   "Carrier_78_SpareSafetyInput(2_3)" AT %I4264.3 : Bool;   // SPARE SAFETY INPUT
   "Carrier_78_SpareSafetyInput(2_4)" AT %I4264.4 : Bool;   // SPARE SAFETY INPUT
   "Carrier_78_SpareSafetyInput(2_5)" AT %I4264.5 : Bool;   // SPARE SAFETY INPUT
   "Carrier_78_SpareSafetyInput(2_6)" AT %I4264.6 : Bool;   // SPARE SAFETY INPUT
   "Carrier_78_SpareSafetyInput(2_7)" AT %I4264.7 : Bool;   // SPARE SAFETY INPUT
   "Carrier_78_Slot3_SafetyOutput" AT %IW4265 : Word;   // SLOT 3 SAFETY OUTPUT WORD
   "Carrier_78_Crash_Detect_OK" AT %I4265.0 : Bool;   // CARRIER CRASH DETECT
   "Carrier_78_SpareSafetyOutput(3_1)" AT %I4265.1 : Bool;   // SPARE SAFETY OUTPUT
   "Carrier_78_SpareSafetyOutput(3_2)" AT %I4265.2 : Bool;   // SPARE SAFETY OUTPUT
   "Carrier_78_SpareSafetyOutput(3_3)" AT %I4265.3 : Bool;   // SPARE SAFETY OUTPUT
   "Carrier_78_SpareSafetyOutput(3_4)" AT %I4265.4 : Bool;   // SPARE SAFETY OUTPUT
   "Carrier_78_SpareSafetyOutput(3_5)" AT %I4265.5 : Bool;   // SPARE SAFETY OUTPUT
   "Carrier_78_SpareSafetyOutput(3_6)" AT %I4265.6 : Bool;   // SPARE SAFETY OUTPUT
   "Carrier_78_SpareSafetyOutput(3_7)" AT %I4265.7 : Bool;   // SPARE SAFETY OUTPUT
   "Carrier_78_Slot4_Input" AT %IW4266 : Word;   // SLOT 4 INPUT WORD
   "Carrier_78_480VPowerOn_MDCB1" AT %I4266.0 : Bool;   // 480 VAC POWER ON MDCB 1
   "Carrier_78_SpareInput(4_1)" AT %I4266.1 : Bool;   // SPARE INPUT
   "Carrier_78_SpareInput(4_2)" AT %I4266.2 : Bool;   // SPARE INPUT
   "Carrier_78_SitopSelectStatus" AT %I4266.3 : Bool;   // SITOP SELECT STATUS
   "Carrier_78_DCsupplyOnPSCB2" AT %I4266.4 : Bool;   // DC SUPPLY ON PSCB 2
   "Carrier_78_SpareInput(4_5)" AT %I4266.5 : Bool;   // SPARE INPUT
   "Carrier_78_SpareInput(4_6)" AT %I4266.6 : Bool;   // SPARE INPUT
   "Carrier_78_SpareInput(4_7)" AT %I4266.7 : Bool;   // SPARE INPUT
   "Carrier_78_PB1_ProdHoldLH" AT %I4267.0 : Bool;   // PB 1 PRODUCTION HOLD LH
   "Carrier_78_PB2_ResetLH" AT %I4267.1 : Bool;   // PB 2 RESET LH
   "Carrier_78_PB3_ProdHoldRH" AT %I4267.2 : Bool;   // PB 3 PRODUCTION HOLD RH
   "Carrier_78_PB4_ResetRH" AT %I4267.3 : Bool;   // PB 4 RESET RH
   "Carrier_78_SpareInput(4_14)" AT %I4267.4 : Bool;   // SPARE INPUT
   "Carrier_78_SpareInput(4_15)" AT %I4267.5 : Bool;   // SPARE INPUT
   "Carrier_78_SpareInput(4_16)" AT %I4267.6 : Bool;   // SPARE INPUT
   "Carrier_78_SpareInput(4_17)" AT %I4267.7 : Bool;   // SPARE INPUT
   "Carrier_78_Slot5_Output" AT %IW4268 : Word;   // SLOT 5 OUTPUT WORD
   "Carrier_78_IRD400_HMI_24VDC_ENABLE" AT %I4268.0 : Bool;   // IRD 400 PANEL HMI 24V DC POWER
   "Carrier_78_FaultLight_LH" AT %I4268.1 : Bool;   // FAULT LIGHT LH
   "Carrier_78_RunLight_LH" AT %I4268.2 : Bool;   // RUN LIGHT LH
   "Carrier_78_FaultLight_RH" AT %I4268.3 : Bool;   // FAULT LIGHT RH
   "Carrier_78_RunLight_RH" AT %I4268.4 : Bool;   // RUN LIGHT RH
   "Carrier_78_SpareOutput(5_5)" AT %I4268.5 : Bool;   // SPARE OUTPUT
   "Carrier_78_SpareOutput(5_6)" AT %I4268.6 : Bool;   // SPARE OUTPUT
   "Carrier_78_SpareOutput(5_7)" AT %I4268.7 : Bool;   // SPARE OUTPUT
   "Carrier_78_ActualSpeed" AT %IW4270 : Word;   // ACTUAL SPEED
   "Carrier_78_CarrierDriveAlarm" AT %IW4272 : Word;   // CARRIER DRIVE ALARM
   "Carrier_78_CarrierDriveWarning" AT %IW4274 : Word;   // CARRIER DRIVE WARNING
   "Carrier_79_Status" AT %IW4300 : Word;   // CARRIER STATUS WORD
   "Carrier_79_Status.0" AT %I4300.0 : Bool;   // HEARTBEAT
   "Carrier_79_Status.1" AT %I4300.1 : Bool;   // MANUAL
   "Carrier_79_Status.2" AT %I4300.2 : Bool;   // IN_AUTO
   "Carrier_79_Status.3" AT %I4300.3 : Bool;   // POSITIONING_COMPLETE
   "Carrier_79_Status.4" AT %I4300.4 : Bool;   // PRODUCTION HOLD
   "Carrier_79_Status.5" AT %I4300.5 : Bool;   // CARRIER MOVING FORWARD
   "Carrier_79_Status.6" AT %I4300.6 : Bool;   // CARRIER MOVING REVERSE
   "Carrier_79_Status.7" AT %I4300.7 : Bool;   // CARRIER FAULT
   "Carrier_79_Status.8" AT %I4301.0 : Bool;   // CRASH DETECT TRIPPED
   "Carrier_79_Status.9" AT %I4301.1 : Bool;
   "Carrier_79_Status.10" AT %I4301.2 : Bool;
   "Carrier_79_Status.11" AT %I4301.3 : Bool;
   "Carrier_79_Status.12" AT %I4301.4 : Bool;
   "Carrier_79_Status.13" AT %I4301.5 : Bool;
   "Carrier_79_Status.14" AT %I4301.6 : Bool;
   "Carrier_79_Status.15" AT %I4301.7 : Bool;
   "Carrier_79_SDCFaultCode" AT %IW4302 : Word;   // SDC FAULT CODE
   "Carrier_79_CarrierPosition" AT %ID4304 : DWord;   // CARRIER POSITION
   "Carrier_79_CarrierNumber" AT %IW4308 : Word;   // CARRIER NUMBER
   "Carrier_79_G120DControlWord" AT %IW4310 : Word;   // G120D_STW1_CONTROL
   "Carrier_79_G120DControlWord.0" AT %I4310.0 : Bool;   // Bit_00_ON
   "Carrier_79_G120DControlWord.1" AT %I4310.1 : Bool;   // Bit_01_AUS2_INH
   "Carrier_79_G120DControlWord.2" AT %I4310.2 : Bool;   // Bit_02_AUS3_STOP
   "Carrier_79_G120DControlWord.3" AT %I4310.3 : Bool;   // Bit_03_EN
   "Carrier_79_G120DControlWord.4" AT %I4310.4 : Bool;   // Bit_04_EN_RAMP
   "Carrier_79_G120DControlWord.5" AT %I4310.5 : Bool;   // Bit_05_START_RAMP
   "Carrier_79_G120DControlWord.6" AT %I4310.6 : Bool;   // Bit_06_SETPOINT
   "Carrier_79_G120DControlWord.7" AT %I4310.7 : Bool;   // Bit_07_RESET
   "Carrier_79_G120DControlWord.8" AT %I4311.0 : Bool;   // Bit_08_JOG_R
   "Carrier_79_G120DControlWord.9" AT %I4311.1 : Bool;   // Bit_09_JOG_L
   "Carrier_79_G120DControlWord.10" AT %I4311.2 : Bool;   // Bit_10_CONTR_PLC
   "Carrier_79_G120DControlWord.11" AT %I4311.3 : Bool;   // Bit_11_REVERSE
   "Carrier_79_G120DControlWord.12" AT %I4311.4 : Bool;   // Bit_12_BRAKE_RELEASE
   "Carrier_79_G120DControlWord.13" AT %I4311.5 : Bool;   // Bit_13_DDS
   "Carrier_79_G120DControlWord.14" AT %I4311.6 : Bool;   // Bit_14_DO0
   "Carrier_79_G120DControlWord.15" AT %I4311.7 : Bool;   // Bit_15_DO1
   "Carrier_79_G120DStatusWord" AT %IW4312 : Word;   // G120D_ZSW1_STATUS
   "Carrier_79_G120DStatusWord.0" AT %I4312.0 : Bool;   // Bit_00_READY_RUN
   "Carrier_79_G120DStatusWord.1" AT %I4312.1 : Bool;   // Bit_01_READY_ON
   "Carrier_79_G120DStatusWord.2" AT %I4312.2 : Bool;   // Bit_02_ENABLE
   "Carrier_79_G120DStatusWord.3" AT %I4312.3 : Bool;   // Bit_03_FAULT
   "Carrier_79_G120DStatusWord.4" AT %I4312.4 : Bool;   // Bit_04_OFF2
   "Carrier_79_G120DStatusWord.5" AT %I4312.5 : Bool;   // Bit_05_OFF3
   "Carrier_79_G120DStatusWord.6" AT %I4312.6 : Bool;   // Bit_06_LOCK_OUT
   "Carrier_79_G120DStatusWord.7" AT %I4312.7 : Bool;   // Bit_07_WARN
   "Carrier_79_G120DStatusWord.8" AT %I4313.0 : Bool;   // Bit_08_NO_DEVIATION
   "Carrier_79_G120DStatusWord.9" AT %I4313.1 : Bool;   // Bit_09_CONTR_PLC
   "Carrier_79_G120DStatusWord.10" AT %I4313.2 : Bool;   // Bit_10_F_MAX
   "Carrier_79_G120DStatusWord.11" AT %I4313.3 : Bool;   // Bit_11_LIMIT_REACHED
   "Carrier_79_G120DStatusWord.12" AT %I4313.4 : Bool;   // Bit_12_BRAKE_OPEN
   "Carrier_79_G120DStatusWord.13" AT %I4313.5 : Bool;   // Bit_13_NO_OVERTEMP
   "Carrier_79_G120DStatusWord.14" AT %I4313.6 : Bool;   // Bit_14_CW_CCW
   "Carrier_79_G120DStatusWord.15" AT %I4313.7 : Bool;   // Bit_15_OVERL
   "Carrier_79_Slot2_Input" AT %IW4314 : Word;   // SLOT 2 INPUT WORD
   "Carrier_79_CrashDetectSW" AT %I4314.0 : Bool;   // CRASH DETECT SW
   "Carrier_79_SpareSafetyInput(2_1)" AT %I4314.1 : Bool;   // SPARE SAFETY INPUT
   "Carrier_79_SpareSafetyInput(2_2)" AT %I4314.2 : Bool;   // SPARE SAFETY INPUT
   "Carrier_79_SpareSafetyInput(2_3)" AT %I4314.3 : Bool;   // SPARE SAFETY INPUT
   "Carrier_79_SpareSafetyInput(2_4)" AT %I4314.4 : Bool;   // SPARE SAFETY INPUT
   "Carrier_79_SpareSafetyInput(2_5)" AT %I4314.5 : Bool;   // SPARE SAFETY INPUT
   "Carrier_79_SpareSafetyInput(2_6)" AT %I4314.6 : Bool;   // SPARE SAFETY INPUT
   "Carrier_79_SpareSafetyInput(2_7)" AT %I4314.7 : Bool;   // SPARE SAFETY INPUT
   "Carrier_79_Slot3_SafetyOutput" AT %IW4315 : Word;   // SLOT 3 SAFETY OUTPUT WORD
   "Carrier_79_Crash_Detect_OK" AT %I4315.0 : Bool;   // CARRIER CRASH DETECT
   "Carrier_79_SpareSafetyOutput(3_1)" AT %I4315.1 : Bool;   // SPARE SAFETY OUTPUT
   "Carrier_79_SpareSafetyOutput(3_2)" AT %I4315.2 : Bool;   // SPARE SAFETY OUTPUT
   "Carrier_79_SpareSafetyOutput(3_3)" AT %I4315.3 : Bool;   // SPARE SAFETY OUTPUT
   "Carrier_79_SpareSafetyOutput(3_4)" AT %I4315.4 : Bool;   // SPARE SAFETY OUTPUT
   "Carrier_79_SpareSafetyOutput(3_5)" AT %I4315.5 : Bool;   // SPARE SAFETY OUTPUT
   "Carrier_79_SpareSafetyOutput(3_6)" AT %I4315.6 : Bool;   // SPARE SAFETY OUTPUT
   "Carrier_79_SpareSafetyOutput(3_7)" AT %I4315.7 : Bool;   // SPARE SAFETY OUTPUT
   "Carrier_79_Slot4_Input" AT %IW4316 : Word;   // SLOT 4 INPUT WORD
   "Carrier_79_480VPowerOn_MDCB1" AT %I4316.0 : Bool;   // 480 VAC POWER ON MDCB 1
   "Carrier_79_SpareInput(4_1)" AT %I4316.1 : Bool;   // SPARE INPUT
   "Carrier_79_SpareInput(4_2)" AT %I4316.2 : Bool;   // SPARE INPUT
   "Carrier_79_SitopSelectStatus" AT %I4316.3 : Bool;   // SITOP SELECT STATUS
   "Carrier_79_DCsupplyOnPSCB2" AT %I4316.4 : Bool;   // DC SUPPLY ON PSCB 2
   "Carrier_79_SpareInput(4_5)" AT %I4316.5 : Bool;   // SPARE INPUT
   "Carrier_79_SpareInput(4_6)" AT %I4316.6 : Bool;   // SPARE INPUT
   "Carrier_79_SpareInput(4_7)" AT %I4316.7 : Bool;   // SPARE INPUT
   "Carrier_79_PB1_ProdHoldLH" AT %I4317.0 : Bool;   // PB 1 PRODUCTION HOLD LH
   "Carrier_79_PB2_ResetLH" AT %I4317.1 : Bool;   // PB 2 RESET LH
   "Carrier_79_PB3_ProdHoldRH" AT %I4317.2 : Bool;   // PB 3 PRODUCTION HOLD RH
   "Carrier_79_PB4_ResetRH" AT %I4317.3 : Bool;   // PB 4 RESET RH
   "Carrier_79_SpareInput(4_14)" AT %I4317.4 : Bool;   // SPARE INPUT
   "Carrier_79_SpareInput(4_15)" AT %I4317.5 : Bool;   // SPARE INPUT
   "Carrier_79_SpareInput(4_16)" AT %I4317.6 : Bool;   // SPARE INPUT
   "Carrier_79_SpareInput(4_17)" AT %I4317.7 : Bool;   // SPARE INPUT
   "Carrier_79_Slot5_Output" AT %IW4318 : Word;   // SLOT 5 OUTPUT WORD
   "Carrier_79_IRD400_HMI_24VDC_ENABLE" AT %I4318.0 : Bool;   // IRD 400 PANEL HMI 24V DC POWER
   "Carrier_79_FaultLight_LH" AT %I4318.1 : Bool;   // FAULT LIGHT LH
   "Carrier_79_RunLight_LH" AT %I4318.2 : Bool;   // RUN LIGHT LH
   "Carrier_79_FaultLight_RH" AT %I4318.3 : Bool;   // FAULT LIGHT RH
   "Carrier_79_RunLight_RH" AT %I4318.4 : Bool;   // RUN LIGHT RH
   "Carrier_79_SpareOutput(5_5)" AT %I4318.5 : Bool;   // SPARE OUTPUT
   "Carrier_79_SpareOutput(5_6)" AT %I4318.6 : Bool;   // SPARE OUTPUT
   "Carrier_79_SpareOutput(5_7)" AT %I4318.7 : Bool;   // SPARE OUTPUT
   "Carrier_79_ActualSpeed" AT %IW4320 : Word;   // ACTUAL SPEED
   "Carrier_79_CarrierDriveAlarm" AT %IW4322 : Word;   // CARRIER DRIVE ALARM
   "Carrier_79_CarrierDriveWarning" AT %IW4324 : Word;   // CARRIER DRIVE WARNING
   "Carrier_80_Status" AT %IW4350 : Word;   // CARRIER STATUS WORD
   "Carrier_80_Status.0" AT %I4350.0 : Bool;   // HEARTBEAT
   "Carrier_80_Status.1" AT %I4350.1 : Bool;   // MANUAL
   "Carrier_80_Status.2" AT %I4350.2 : Bool;   // IN_AUTO
   "Carrier_80_Status.3" AT %I4350.3 : Bool;   // POSITIONING_COMPLETE
   "Carrier_80_Status.4" AT %I4350.4 : Bool;   // PRODUCTION HOLD
   "Carrier_80_Status.5" AT %I4350.5 : Bool;   // CARRIER MOVING FORWARD
   "Carrier_80_Status.6" AT %I4350.6 : Bool;   // CARRIER MOVING REVERSE
   "Carrier_80_Status.7" AT %I4350.7 : Bool;   // CARRIER FAULT
   "Carrier_80_Status.8" AT %I4351.0 : Bool;   // CRASH DETECT TRIPPED
   "Carrier_80_Status.9" AT %I4351.1 : Bool;
   "Carrier_80_Status.10" AT %I4351.2 : Bool;
   "Carrier_80_Status.11" AT %I4351.3 : Bool;
   "Carrier_80_Status.12" AT %I4351.4 : Bool;
   "Carrier_80_Status.13" AT %I4351.5 : Bool;
   "Carrier_80_Status.14" AT %I4351.6 : Bool;
   "Carrier_80_Status.15" AT %I4351.7 : Bool;
   "Carrier_80_SDCFaultCode" AT %IW4352 : Word;   // SDC FAULT CODE
   "Carrier_80_CarrierPosition" AT %ID4354 : DWord;   // CARRIER POSITION
   "Carrier_80_CarrierNumber" AT %IW4358 : Word;   // CARRIER NUMBER
   "Carrier_80_G120DControlWord" AT %IW4360 : Word;   // G120D_STW1_CONTROL
   "Carrier_80_G120DControlWord.0" AT %I4360.0 : Bool;   // Bit_00_ON
   "Carrier_80_G120DControlWord.1" AT %I4360.1 : Bool;   // Bit_01_AUS2_INH
   "Carrier_80_G120DControlWord.2" AT %I4360.2 : Bool;   // Bit_02_AUS3_STOP
   "Carrier_80_G120DControlWord.3" AT %I4360.3 : Bool;   // Bit_03_EN
   "Carrier_80_G120DControlWord.4" AT %I4360.4 : Bool;   // Bit_04_EN_RAMP
   "Carrier_80_G120DControlWord.5" AT %I4360.5 : Bool;   // Bit_05_START_RAMP
   "Carrier_80_G120DControlWord.6" AT %I4360.6 : Bool;   // Bit_06_SETPOINT
   "Carrier_80_G120DControlWord.7" AT %I4360.7 : Bool;   // Bit_07_RESET
   "Carrier_80_G120DControlWord.8" AT %I4361.0 : Bool;   // Bit_08_JOG_R
   "Carrier_80_G120DControlWord.9" AT %I4361.1 : Bool;   // Bit_09_JOG_L
   "Carrier_80_G120DControlWord.10" AT %I4361.2 : Bool;   // Bit_10_CONTR_PLC
   "Carrier_80_G120DControlWord.11" AT %I4361.3 : Bool;   // Bit_11_REVERSE
   "Carrier_80_G120DControlWord.12" AT %I4361.4 : Bool;   // Bit_12_BRAKE_RELEASE
   "Carrier_80_G120DControlWord.13" AT %I4361.5 : Bool;   // Bit_13_DDS
   "Carrier_80_G120DControlWord.14" AT %I4361.6 : Bool;   // Bit_14_DO0
   "Carrier_80_G120DControlWord.15" AT %I4361.7 : Bool;   // Bit_15_DO1
   "Carrier_80_G120DStatusWord" AT %IW4362 : Word;   // G120D_ZSW1_STATUS
   "Carrier_80_G120DStatusWord.0" AT %I4362.0 : Bool;   // Bit_00_READY_RUN
   "Carrier_80_G120DStatusWord.1" AT %I4362.1 : Bool;   // Bit_01_READY_ON
   "Carrier_80_G120DStatusWord.2" AT %I4362.2 : Bool;   // Bit_02_ENABLE
   "Carrier_80_G120DStatusWord.3" AT %I4362.3 : Bool;   // Bit_03_FAULT
   "Carrier_80_G120DStatusWord.4" AT %I4362.4 : Bool;   // Bit_04_OFF2
   "Carrier_80_G120DStatusWord.5" AT %I4362.5 : Bool;   // Bit_05_OFF3
   "Carrier_80_G120DStatusWord.6" AT %I4362.6 : Bool;   // Bit_06_LOCK_OUT
   "Carrier_80_G120DStatusWord.7" AT %I4362.7 : Bool;   // Bit_07_WARN
   "Carrier_80_G120DStatusWord.8" AT %I4363.0 : Bool;   // Bit_08_NO_DEVIATION
   "Carrier_80_G120DStatusWord.9" AT %I4363.1 : Bool;   // Bit_09_CONTR_PLC
   "Carrier_80_G120DStatusWord.10" AT %I4363.2 : Bool;   // Bit_10_F_MAX
   "Carrier_80_G120DStatusWord.11" AT %I4363.3 : Bool;   // Bit_11_LIMIT_REACHED
   "Carrier_80_G120DStatusWord.12" AT %I4363.4 : Bool;   // Bit_12_BRAKE_OPEN
   "Carrier_80_G120DStatusWord.13" AT %I4363.5 : Bool;   // Bit_13_NO_OVERTEMP
   "Carrier_80_G120DStatusWord.14" AT %I4363.6 : Bool;   // Bit_14_CW_CCW
   "Carrier_80_G120DStatusWord.15" AT %I4363.7 : Bool;   // Bit_15_OVERL
   "Carrier_80_Slot2_Input" AT %IW4364 : Word;   // SLOT 2 INPUT WORD
   "Carrier_80_CrashDetectSW" AT %I4364.0 : Bool;   // CRASH DETECT SW
   "Carrier_80_SpareSafetyInput(2_1)" AT %I4364.1 : Bool;   // SPARE SAFETY INPUT
   "Carrier_80_SpareSafetyInput(2_2)" AT %I4364.2 : Bool;   // SPARE SAFETY INPUT
   "Carrier_80_SpareSafetyInput(2_3)" AT %I4364.3 : Bool;   // SPARE SAFETY INPUT
   "Carrier_80_SpareSafetyInput(2_4)" AT %I4364.4 : Bool;   // SPARE SAFETY INPUT
   "Carrier_80_SpareSafetyInput(2_5)" AT %I4364.5 : Bool;   // SPARE SAFETY INPUT
   "Carrier_80_SpareSafetyInput(2_6)" AT %I4364.6 : Bool;   // SPARE SAFETY INPUT
   "Carrier_80_SpareSafetyInput(2_7)" AT %I4364.7 : Bool;   // SPARE SAFETY INPUT
   "Carrier_80_Slot3_SafetyOutput" AT %IW4365 : Word;   // SLOT 3 SAFETY OUTPUT WORD
   "Carrier_80_Crash_Detect_OK" AT %I4365.0 : Bool;   // CARRIER CRASH DETECT
   "Carrier_80_SpareSafetyOutput(3_1)" AT %I4365.1 : Bool;   // SPARE SAFETY OUTPUT
   "Carrier_80_SpareSafetyOutput(3_2)" AT %I4365.2 : Bool;   // SPARE SAFETY OUTPUT
   "Carrier_80_SpareSafetyOutput(3_3)" AT %I4365.3 : Bool;   // SPARE SAFETY OUTPUT
   "Carrier_80_SpareSafetyOutput(3_4)" AT %I4365.4 : Bool;   // SPARE SAFETY OUTPUT
   "Carrier_80_SpareSafetyOutput(3_5)" AT %I4365.5 : Bool;   // SPARE SAFETY OUTPUT
   "Carrier_80_SpareSafetyOutput(3_6)" AT %I4365.6 : Bool;   // SPARE SAFETY OUTPUT
   "Carrier_80_SpareSafetyOutput(3_7)" AT %I4365.7 : Bool;   // SPARE SAFETY OUTPUT
   "Carrier_80_Slot4_Input" AT %IW4366 : Word;   // SLOT 4 INPUT WORD
   "Carrier_80_480VPowerOn_MDCB1" AT %I4366.0 : Bool;   // 480 VAC POWER ON MDCB 1
   "Carrier_80_SpareInput(4_1)" AT %I4366.1 : Bool;   // SPARE INPUT
   "Carrier_80_SpareInput(4_2)" AT %I4366.2 : Bool;   // SPARE INPUT
   "Carrier_80_SitopSelectStatus" AT %I4366.3 : Bool;   // SITOP SELECT STATUS
   "Carrier_80_DCsupplyOnPSCB2" AT %I4366.4 : Bool;   // DC SUPPLY ON PSCB 2
   "Carrier_80_SpareInput(4_5)" AT %I4366.5 : Bool;   // SPARE INPUT
   "Carrier_80_SpareInput(4_6)" AT %I4366.6 : Bool;   // SPARE INPUT
   "Carrier_80_SpareInput(4_7)" AT %I4366.7 : Bool;   // SPARE INPUT
   "Carrier_80_PB1_ProdHoldLH" AT %I4367.0 : Bool;   // PB 1 PRODUCTION HOLD LH
   "Carrier_80_PB2_ResetLH" AT %I4367.1 : Bool;   // PB 2 RESET LH
   "Carrier_80_PB3_ProdHoldRH" AT %I4367.2 : Bool;   // PB 3 PRODUCTION HOLD RH
   "Carrier_80_PB4_ResetRH" AT %I4367.3 : Bool;   // PB 4 RESET RH
   "Carrier_80_SpareInput(4_14)" AT %I4367.4 : Bool;   // SPARE INPUT
   "Carrier_80_SpareInput(4_15)" AT %I4367.5 : Bool;   // SPARE INPUT
   "Carrier_80_SpareInput(4_16)" AT %I4367.6 : Bool;   // SPARE INPUT
   "Carrier_80_SpareInput(4_17)" AT %I4367.7 : Bool;   // SPARE INPUT
   "Carrier_80_Slot5_Output" AT %IW4368 : Word;   // SLOT 5 OUTPUT WORD
   "Carrier_80_IRD400_HMI_24VDC_ENABLE" AT %I4368.0 : Bool;   // IRD 400 PANEL HMI 24V DC POWER
   "Carrier_80_FaultLight_LH" AT %I4368.1 : Bool;   // FAULT LIGHT LH
   "Carrier_80_RunLight_LH" AT %I4368.2 : Bool;   // RUN LIGHT LH
   "Carrier_80_FaultLight_RH" AT %I4368.3 : Bool;   // FAULT LIGHT RH
   "Carrier_80_RunLight_RH" AT %I4368.4 : Bool;   // RUN LIGHT RH
   "Carrier_80_SpareOutput(5_5)" AT %I4368.5 : Bool;   // SPARE OUTPUT
   "Carrier_80_SpareOutput(5_6)" AT %I4368.6 : Bool;   // SPARE OUTPUT
   "Carrier_80_SpareOutput(5_7)" AT %I4368.7 : Bool;   // SPARE OUTPUT
   "Carrier_80_ActualSpeed" AT %IW4370 : Word;   // ACTUAL SPEED
   "Carrier_80_CarrierDriveAlarm" AT %IW4372 : Word;   // CARRIER DRIVE ALARM
   "Carrier_80_CarrierDriveWarning" AT %IW4374 : Word;   // CARRIER DRIVE WARNING
   "Carrier_81_Status" AT %IW4400 : Word;   // CARRIER STATUS WORD
   "Carrier_81_Status.0" AT %I4400.0 : Bool;   // HEARTBEAT
   "Carrier_81_Status.1" AT %I4400.1 : Bool;   // MANUAL
   "Carrier_81_Status.2" AT %I4400.2 : Bool;   // IN_AUTO
   "Carrier_81_Status.3" AT %I4400.3 : Bool;   // POSITIONING_COMPLETE
   "Carrier_81_Status.4" AT %I4400.4 : Bool;   // PRODUCTION HOLD
   "Carrier_81_Status.5" AT %I4400.5 : Bool;   // CARRIER MOVING FORWARD
   "Carrier_81_Status.6" AT %I4400.6 : Bool;   // CARRIER MOVING REVERSE
   "Carrier_81_Status.7" AT %I4400.7 : Bool;   // CARRIER FAULT
   "Carrier_81_Status.8" AT %I4401.0 : Bool;   // CRASH DETECT TRIPPED
   "Carrier_81_Status.9" AT %I4401.1 : Bool;
   "Carrier_81_Status.10" AT %I4401.2 : Bool;
   "Carrier_81_Status.11" AT %I4401.3 : Bool;
   "Carrier_81_Status.12" AT %I4401.4 : Bool;
   "Carrier_81_Status.13" AT %I4401.5 : Bool;
   "Carrier_81_Status.14" AT %I4401.6 : Bool;
   "Carrier_81_Status.15" AT %I4401.7 : Bool;
   "Carrier_81_SDCFaultCode" AT %IW4402 : Word;   // SDC FAULT CODE
   "Carrier_81_CarrierPosition" AT %ID4404 : DWord;   // CARRIER POSITION
   "Carrier_81_CarrierNumber" AT %IW4408 : Word;   // CARRIER NUMBER
   "Carrier_81_G120DControlWord" AT %IW4410 : Word;   // G120D_STW1_CONTROL
   "Carrier_81_G120DControlWord.0" AT %I4410.0 : Bool;   // Bit_00_ON
   "Carrier_81_G120DControlWord.1" AT %I4410.1 : Bool;   // Bit_01_AUS2_INH
   "Carrier_81_G120DControlWord.2" AT %I4410.2 : Bool;   // Bit_02_AUS3_STOP
   "Carrier_81_G120DControlWord.3" AT %I4410.3 : Bool;   // Bit_03_EN
   "Carrier_81_G120DControlWord.4" AT %I4410.4 : Bool;   // Bit_04_EN_RAMP
   "Carrier_81_G120DControlWord.5" AT %I4410.5 : Bool;   // Bit_05_START_RAMP
   "Carrier_81_G120DControlWord.6" AT %I4410.6 : Bool;   // Bit_06_SETPOINT
   "Carrier_81_G120DControlWord.7" AT %I4410.7 : Bool;   // Bit_07_RESET
   "Carrier_81_G120DControlWord.8" AT %I4411.0 : Bool;   // Bit_08_JOG_R
   "Carrier_81_G120DControlWord.9" AT %I4411.1 : Bool;   // Bit_09_JOG_L
   "Carrier_81_G120DControlWord.10" AT %I4411.2 : Bool;   // Bit_10_CONTR_PLC
   "Carrier_81_G120DControlWord.11" AT %I4411.3 : Bool;   // Bit_11_REVERSE
   "Carrier_81_G120DControlWord.12" AT %I4411.4 : Bool;   // Bit_12_BRAKE_RELEASE
   "Carrier_81_G120DControlWord.13" AT %I4411.5 : Bool;   // Bit_13_DDS
   "Carrier_81_G120DControlWord.14" AT %I4411.6 : Bool;   // Bit_14_DO0
   "Carrier_81_G120DControlWord.15" AT %I4411.7 : Bool;   // Bit_15_DO1
   "Carrier_81_G120DStatusWord" AT %IW4412 : Word;   // G120D_ZSW1_STATUS
   "Carrier_81_G120DStatusWord.0" AT %I4412.0 : Bool;   // Bit_00_READY_RUN
   "Carrier_81_G120DStatusWord.1" AT %I4412.1 : Bool;   // Bit_01_READY_ON
   "Carrier_81_G120DStatusWord.2" AT %I4412.2 : Bool;   // Bit_02_ENABLE
   "Carrier_81_G120DStatusWord.3" AT %I4412.3 : Bool;   // Bit_03_FAULT
   "Carrier_81_G120DStatusWord.4" AT %I4412.4 : Bool;   // Bit_04_OFF2
   "Carrier_81_G120DStatusWord.5" AT %I4412.5 : Bool;   // Bit_05_OFF3
   "Carrier_81_G120DStatusWord.6" AT %I4412.6 : Bool;   // Bit_06_LOCK_OUT
   "Carrier_81_G120DStatusWord.7" AT %I4412.7 : Bool;   // Bit_07_WARN
   "Carrier_81_G120DStatusWord.8" AT %I4413.0 : Bool;   // Bit_08_NO_DEVIATION
   "Carrier_81_G120DStatusWord.9" AT %I4413.1 : Bool;   // Bit_09_CONTR_PLC
   "Carrier_81_G120DStatusWord.10" AT %I4413.2 : Bool;   // Bit_10_F_MAX
   "Carrier_81_G120DStatusWord.11" AT %I4413.3 : Bool;   // Bit_11_LIMIT_REACHED
   "Carrier_81_G120DStatusWord.12" AT %I4413.4 : Bool;   // Bit_12_BRAKE_OPEN
   "Carrier_81_G120DStatusWord.13" AT %I4413.5 : Bool;   // Bit_13_NO_OVERTEMP
   "Carrier_81_G120DStatusWord.14" AT %I4413.6 : Bool;   // Bit_14_CW_CCW
   "Carrier_81_G120DStatusWord.15" AT %I4413.7 : Bool;   // Bit_15_OVERL
   "Carrier_81_Slot2_Input" AT %IW4414 : Word;   // SLOT 2 INPUT WORD
   "Carrier_81_CrashDetectSW" AT %I4414.0 : Bool;   // CRASH DETECT SW
   "Carrier_81_SpareSafetyInput(2_1)" AT %I4414.1 : Bool;   // SPARE SAFETY INPUT
   "Carrier_81_SpareSafetyInput(2_2)" AT %I4414.2 : Bool;   // SPARE SAFETY INPUT
   "Carrier_81_SpareSafetyInput(2_3)" AT %I4414.3 : Bool;   // SPARE SAFETY INPUT
   "Carrier_81_SpareSafetyInput(2_4)" AT %I4414.4 : Bool;   // SPARE SAFETY INPUT
   "Carrier_81_SpareSafetyInput(2_5)" AT %I4414.5 : Bool;   // SPARE SAFETY INPUT
   "Carrier_81_SpareSafetyInput(2_6)" AT %I4414.6 : Bool;   // SPARE SAFETY INPUT
   "Carrier_81_SpareSafetyInput(2_7)" AT %I4414.7 : Bool;   // SPARE SAFETY INPUT
   "Carrier_81_Slot3_SafetyOutput" AT %IW4415 : Word;   // SLOT 3 SAFETY OUTPUT WORD
   "Carrier_81_Crash_Detect_OK" AT %I4415.0 : Bool;   // CARRIER CRASH DETECT
   "Carrier_81_SpareSafetyOutput(3_1)" AT %I4415.1 : Bool;   // SPARE SAFETY OUTPUT
   "Carrier_81_SpareSafetyOutput(3_2)" AT %I4415.2 : Bool;   // SPARE SAFETY OUTPUT
   "Carrier_81_SpareSafetyOutput(3_3)" AT %I4415.3 : Bool;   // SPARE SAFETY OUTPUT
   "Carrier_81_SpareSafetyOutput(3_4)" AT %I4415.4 : Bool;   // SPARE SAFETY OUTPUT
   "Carrier_81_SpareSafetyOutput(3_5)" AT %I4415.5 : Bool;   // SPARE SAFETY OUTPUT
   "Carrier_81_SpareSafetyOutput(3_6)" AT %I4415.6 : Bool;   // SPARE SAFETY OUTPUT
   "Carrier_81_SpareSafetyOutput(3_7)" AT %I4415.7 : Bool;   // SPARE SAFETY OUTPUT
   "Carrier_81_Slot4_Input" AT %IW4416 : Word;   // SLOT 4 INPUT WORD
   "Carrier_81_480VPowerOn_MDCB1" AT %I4416.0 : Bool;   // 480 VAC POWER ON MDCB 1
   "Carrier_81_SpareInput(4_1)" AT %I4416.1 : Bool;   // SPARE INPUT
   "Carrier_81_SpareInput(4_2)" AT %I4416.2 : Bool;   // SPARE INPUT
   "Carrier_81_SitopSelectStatus" AT %I4416.3 : Bool;   // SITOP SELECT STATUS
   "Carrier_81_DCsupplyOnPSCB2" AT %I4416.4 : Bool;   // DC SUPPLY ON PSCB 2
   "Carrier_81_SpareInput(4_5)" AT %I4416.5 : Bool;   // SPARE INPUT
   "Carrier_81_SpareInput(4_6)" AT %I4416.6 : Bool;   // SPARE INPUT
   "Carrier_81_SpareInput(4_7)" AT %I4416.7 : Bool;   // SPARE INPUT
   "Carrier_81_PB1_ProdHoldLH" AT %I4417.0 : Bool;   // PB 1 PRODUCTION HOLD LH
   "Carrier_81_PB2_ResetLH" AT %I4417.1 : Bool;   // PB 2 RESET LH
   "Carrier_81_PB3_ProdHoldRH" AT %I4417.2 : Bool;   // PB 3 PRODUCTION HOLD RH
   "Carrier_81_PB4_ResetRH" AT %I4417.3 : Bool;   // PB 4 RESET RH
   "Carrier_81_SpareInput(4_14)" AT %I4417.4 : Bool;   // SPARE INPUT
   "Carrier_81_SpareInput(4_15)" AT %I4417.5 : Bool;   // SPARE INPUT
   "Carrier_81_SpareInput(4_16)" AT %I4417.6 : Bool;   // SPARE INPUT
   "Carrier_81_SpareInput(4_17)" AT %I4417.7 : Bool;   // SPARE INPUT
   "Carrier_81_Slot5_Output" AT %IW4418 : Word;   // SLOT 5 OUTPUT WORD
   "Carrier_81_IRD400_HMI_24VDC_ENABLE" AT %I4418.0 : Bool;   // IRD 400 PANEL HMI 24V DC POWER
   "Carrier_81_FaultLight_LH" AT %I4418.1 : Bool;   // FAULT LIGHT LH
   "Carrier_81_RunLight_LH" AT %I4418.2 : Bool;   // RUN LIGHT LH
   "Carrier_81_FaultLight_RH" AT %I4418.3 : Bool;   // FAULT LIGHT RH
   "Carrier_81_RunLight_RH" AT %I4418.4 : Bool;   // RUN LIGHT RH
   "Carrier_81_SpareOutput(5_5)" AT %I4418.5 : Bool;   // SPARE OUTPUT
   "Carrier_81_SpareOutput(5_6)" AT %I4418.6 : Bool;   // SPARE OUTPUT
   "Carrier_81_SpareOutput(5_7)" AT %I4418.7 : Bool;   // SPARE OUTPUT
   "Carrier_81_ActualSpeed" AT %IW4420 : Word;   // ACTUAL SPEED
   "Carrier_81_CarrierDriveAlarm" AT %IW4422 : Word;   // CARRIER DRIVE ALARM
   "Carrier_81_CarrierDriveWarning" AT %IW4424 : Word;   // CARRIER DRIVE WARNING
   "Carrier_82_Status" AT %IW4450 : Word;   // CARRIER STATUS WORD
   "Carrier_82_Status.0" AT %I4450.0 : Bool;   // HEARTBEAT
   "Carrier_82_Status.1" AT %I4450.1 : Bool;   // MANUAL
   "Carrier_82_Status.2" AT %I4450.2 : Bool;   // IN_AUTO
   "Carrier_82_Status.3" AT %I4450.3 : Bool;   // POSITIONING_COMPLETE
   "Carrier_82_Status.4" AT %I4450.4 : Bool;   // PRODUCTION HOLD
   "Carrier_82_Status.5" AT %I4450.5 : Bool;   // CARRIER MOVING FORWARD
   "Carrier_82_Status.6" AT %I4450.6 : Bool;   // CARRIER MOVING REVERSE
   "Carrier_82_Status.7" AT %I4450.7 : Bool;   // CARRIER FAULT
   "Carrier_82_Status.8" AT %I4451.0 : Bool;   // CRASH DETECT TRIPPED
   "Carrier_82_Status.9" AT %I4451.1 : Bool;
   "Carrier_82_Status.10" AT %I4451.2 : Bool;
   "Carrier_82_Status.11" AT %I4451.3 : Bool;
   "Carrier_82_Status.12" AT %I4451.4 : Bool;
   "Carrier_82_Status.13" AT %I4451.5 : Bool;
   "Carrier_82_Status.14" AT %I4451.6 : Bool;
   "Carrier_82_Status.15" AT %I4451.7 : Bool;
   "Carrier_82_SDCFaultCode" AT %IW4452 : Word;   // SDC FAULT CODE
   "Carrier_82_CarrierPosition" AT %ID4454 : DWord;   // CARRIER POSITION
   "Carrier_82_CarrierNumber" AT %IW4458 : Word;   // CARRIER NUMBER
   "Carrier_82_G120DControlWord" AT %IW4460 : Word;   // G120D_STW1_CONTROL
   "Carrier_82_G120DControlWord.0" AT %I4460.0 : Bool;   // Bit_00_ON
   "Carrier_82_G120DControlWord.1" AT %I4460.1 : Bool;   // Bit_01_AUS2_INH
   "Carrier_82_G120DControlWord.2" AT %I4460.2 : Bool;   // Bit_02_AUS3_STOP
   "Carrier_82_G120DControlWord.3" AT %I4460.3 : Bool;   // Bit_03_EN
   "Carrier_82_G120DControlWord.4" AT %I4460.4 : Bool;   // Bit_04_EN_RAMP
   "Carrier_82_G120DControlWord.5" AT %I4460.5 : Bool;   // Bit_05_START_RAMP
   "Carrier_82_G120DControlWord.6" AT %I4460.6 : Bool;   // Bit_06_SETPOINT
   "Carrier_82_G120DControlWord.7" AT %I4460.7 : Bool;   // Bit_07_RESET
   "Carrier_82_G120DControlWord.8" AT %I4461.0 : Bool;   // Bit_08_JOG_R
   "Carrier_82_G120DControlWord.9" AT %I4461.1 : Bool;   // Bit_09_JOG_L
   "Carrier_82_G120DControlWord.10" AT %I4461.2 : Bool;   // Bit_10_CONTR_PLC
   "Carrier_82_G120DControlWord.11" AT %I4461.3 : Bool;   // Bit_11_REVERSE
   "Carrier_82_G120DControlWord.12" AT %I4461.4 : Bool;   // Bit_12_BRAKE_RELEASE
   "Carrier_82_G120DControlWord.13" AT %I4461.5 : Bool;   // Bit_13_DDS
   "Carrier_82_G120DControlWord.14" AT %I4461.6 : Bool;   // Bit_14_DO0
   "Carrier_82_G120DControlWord.15" AT %I4461.7 : Bool;   // Bit_15_DO1
   "Carrier_82_G120DStatusWord" AT %IW4462 : Word;   // G120D_ZSW1_STATUS
   "Carrier_82_G120DStatusWord.0" AT %I4462.0 : Bool;   // Bit_00_READY_RUN
   "Carrier_82_G120DStatusWord.1" AT %I4462.1 : Bool;   // Bit_01_READY_ON
   "Carrier_82_G120DStatusWord.2" AT %I4462.2 : Bool;   // Bit_02_ENABLE
   "Carrier_82_G120DStatusWord.3" AT %I4462.3 : Bool;   // Bit_03_FAULT
   "Carrier_82_G120DStatusWord.4" AT %I4462.4 : Bool;   // Bit_04_OFF2
   "Carrier_82_G120DStatusWord.5" AT %I4462.5 : Bool;   // Bit_05_OFF3
   "Carrier_82_G120DStatusWord.6" AT %I4462.6 : Bool;   // Bit_06_LOCK_OUT
   "Carrier_82_G120DStatusWord.7" AT %I4462.7 : Bool;   // Bit_07_WARN
   "Carrier_82_G120DStatusWord.8" AT %I4463.0 : Bool;   // Bit_08_NO_DEVIATION
   "Carrier_82_G120DStatusWord.9" AT %I4463.1 : Bool;   // Bit_09_CONTR_PLC
   "Carrier_82_G120DStatusWord.10" AT %I4463.2 : Bool;   // Bit_10_F_MAX
   "Carrier_82_G120DStatusWord.11" AT %I4463.3 : Bool;   // Bit_11_LIMIT_REACHED
   "Carrier_82_G120DStatusWord.12" AT %I4463.4 : Bool;   // Bit_12_BRAKE_OPEN
   "Carrier_82_G120DStatusWord.13" AT %I4463.5 : Bool;   // Bit_13_NO_OVERTEMP
   "Carrier_82_G120DStatusWord.14" AT %I4463.6 : Bool;   // Bit_14_CW_CCW
   "Carrier_82_G120DStatusWord.15" AT %I4463.7 : Bool;   // Bit_15_OVERL
   "Carrier_82_Slot2_Input" AT %IW4464 : Word;   // SLOT 2 INPUT WORD
   "Carrier_82_CrashDetectSW" AT %I4464.0 : Bool;   // CRASH DETECT SW
   "Carrier_82_SpareSafetyInput(2_1)" AT %I4464.1 : Bool;   // SPARE SAFETY INPUT
   "Carrier_82_SpareSafetyInput(2_2)" AT %I4464.2 : Bool;   // SPARE SAFETY INPUT
   "Carrier_82_SpareSafetyInput(2_3)" AT %I4464.3 : Bool;   // SPARE SAFETY INPUT
   "Carrier_82_SpareSafetyInput(2_4)" AT %I4464.4 : Bool;   // SPARE SAFETY INPUT
   "Carrier_82_SpareSafetyInput(2_5)" AT %I4464.5 : Bool;   // SPARE SAFETY INPUT
   "Carrier_82_SpareSafetyInput(2_6)" AT %I4464.6 : Bool;   // SPARE SAFETY INPUT
   "Carrier_82_SpareSafetyInput(2_7)" AT %I4464.7 : Bool;   // SPARE SAFETY INPUT
   "Carrier_82_Slot3_SafetyOutput" AT %IW4465 : Word;   // SLOT 3 SAFETY OUTPUT WORD
   "Carrier_82_Crash_Detect_OK" AT %I4465.0 : Bool;   // CARRIER CRASH DETECT
   "Carrier_82_SpareSafetyOutput(3_1)" AT %I4465.1 : Bool;   // SPARE SAFETY OUTPUT
   "Carrier_82_SpareSafetyOutput(3_2)" AT %I4465.2 : Bool;   // SPARE SAFETY OUTPUT
   "Carrier_82_SpareSafetyOutput(3_3)" AT %I4465.3 : Bool;   // SPARE SAFETY OUTPUT
   "Carrier_82_SpareSafetyOutput(3_4)" AT %I4465.4 : Bool;   // SPARE SAFETY OUTPUT
   "Carrier_82_SpareSafetyOutput(3_5)" AT %I4465.5 : Bool;   // SPARE SAFETY OUTPUT
   "Carrier_82_SpareSafetyOutput(3_6)" AT %I4465.6 : Bool;   // SPARE SAFETY OUTPUT
   "Carrier_82_SpareSafetyOutput(3_7)" AT %I4465.7 : Bool;   // SPARE SAFETY OUTPUT
   "Carrier_82_Slot4_Input" AT %IW4466 : Word;   // SLOT 4 INPUT WORD
   "Carrier_82_480VPowerOn_MDCB1" AT %I4466.0 : Bool;   // 480 VAC POWER ON MDCB 1
   "Carrier_82_SpareInput(4_1)" AT %I4466.1 : Bool;   // SPARE INPUT
   "Carrier_82_SpareInput(4_2)" AT %I4466.2 : Bool;   // SPARE INPUT
   "Carrier_82_SitopSelectStatus" AT %I4466.3 : Bool;   // SITOP SELECT STATUS
   "Carrier_82_DCsupplyOnPSCB2" AT %I4466.4 : Bool;   // DC SUPPLY ON PSCB 2
   "Carrier_82_SpareInput(4_5)" AT %I4466.5 : Bool;   // SPARE INPUT
   "Carrier_82_SpareInput(4_6)" AT %I4466.6 : Bool;   // SPARE INPUT
   "Carrier_82_SpareInput(4_7)" AT %I4466.7 : Bool;   // SPARE INPUT
   "Carrier_82_PB1_ProdHoldLH" AT %I4467.0 : Bool;   // PB 1 PRODUCTION HOLD LH
   "Carrier_82_PB2_ResetLH" AT %I4467.1 : Bool;   // PB 2 RESET LH
   "Carrier_82_PB3_ProdHoldRH" AT %I4467.2 : Bool;   // PB 3 PRODUCTION HOLD RH
   "Carrier_82_PB4_ResetRH" AT %I4467.3 : Bool;   // PB 4 RESET RH
   "Carrier_82_SpareInput(4_14)" AT %I4467.4 : Bool;   // SPARE INPUT
   "Carrier_82_SpareInput(4_15)" AT %I4467.5 : Bool;   // SPARE INPUT
   "Carrier_82_SpareInput(4_16)" AT %I4467.6 : Bool;   // SPARE INPUT
   "Carrier_82_SpareInput(4_17)" AT %I4467.7 : Bool;   // SPARE INPUT
   "Carrier_82_Slot5_Output" AT %IW4468 : Word;   // SLOT 5 OUTPUT WORD
   "Carrier_82_IRD400_HMI_24VDC_ENABLE" AT %I4468.0 : Bool;   // IRD 400 PANEL HMI 24V DC POWER
   "Carrier_82_FaultLight_LH" AT %I4468.1 : Bool;   // FAULT LIGHT LH
   "Carrier_82_RunLight_LH" AT %I4468.2 : Bool;   // RUN LIGHT LH
   "Carrier_82_FaultLight_RH" AT %I4468.3 : Bool;   // FAULT LIGHT RH
   "Carrier_82_RunLight_RH" AT %I4468.4 : Bool;   // RUN LIGHT RH
   "Carrier_82_SpareOutput(5_5)" AT %I4468.5 : Bool;   // SPARE OUTPUT
   "Carrier_82_SpareOutput(5_6)" AT %I4468.6 : Bool;   // SPARE OUTPUT
   "Carrier_82_SpareOutput(5_7)" AT %I4468.7 : Bool;   // SPARE OUTPUT
   "Carrier_82_ActualSpeed" AT %IW4470 : Word;   // ACTUAL SPEED
   "Carrier_82_CarrierDriveAlarm" AT %IW4472 : Word;   // CARRIER DRIVE ALARM
   "Carrier_82_CarrierDriveWarning" AT %IW4474 : Word;   // CARRIER DRIVE WARNING
   "Tag_101" AT %M2.3 : Bool;
   "Tag_100" AT %M3.7 : Bool;
   "Tag_117" AT %MW58 : Word;
   "SDC_EMS01_Carrier27_Position" AT %QD6104 : DWord;
END_VAR

